screen "Inert Gas Generator Setup" 1280x800, template "Template"
   Circle "Circle_2" at 221,236 size 29x29
      Appearance <- "82_To_HMI_CRNT_MODE_IGG"
   Button "HmiScreenItemData_1" at 1,1 size 150x43; TextOn 'Back'; TextOff 'Main Index'
      on Release: ActivateScreen("02 Main Index", 0)
   Button "HmiScreenItemData_8" at 44,70 size 230x29; TextOn 'Back'; TextOff 'IGGS Mode of Operation'
   Circle "Circle_1" at 221,177 size 29x29
      Appearance <- "82_To_HMI_CRNT_MODE_IGG"
   Button "HmiScreenItemData_4" at 50,167 size 150x51; TextOn 'Back'; TextOff 'Manual'; Authorization "Operate"
      on Press: function_b14e0dd5("80_From_HMI_Request_Manual(1)", 0)
   Circle "Circle_9" at 221,116 size 29x29
      Appearance <- "82_To_HMI_CRNT_MODE_IGG"
   TextField "Text field_1" at 54,547 size 182x20; Text 'Cooling System Overrun'
   TextField "Text field_2" at 54,589 size 192x20; Text 'BWT O2 Content Setpoint'
   TextField "Text field_3" at 54,511 size 89x20; Text 'Description'
   TextField "Text field_5" at 54,670 size 274x20; Text 'IGG Combustion Chamber Post Purge'
   TextField "Text field_6" at 347,511 size 68x20; Text 'Setpoint'
   Button "HmiScreenItemData_6" at 44,467 size 401x29; TextOn 'Back'; TextOff 'IGGS Settings'
   IOField "I/O field_4" at 345,542 size 90x30; Authorization "Commissioning"; FormatPattern 999; Unit  s
      ProcessValue <- "80_From_HMI_Cooling System Overrun"
   IOField "I/O field_5" at 345,583 size 90x30; Authorization "Commissioning"; FormatPattern 99.99; Unit %
      ProcessValue <- "84_Setpoints_E600_BWT_Target"
   IOField "I/O field_6" at 345,664 size 90x30; Authorization "Commissioning"; FormatPattern 999; Unit  s
      ProcessValue <- "80_From_HMI_Post Purge Time"
   TextField "Text field_4" at 54,711 size 294x20; Text 'Air / Inert Gas Pressure (Pre-Ignition)'
   IOField "I/O field_1" at 345,706 size 90x30; Authorization "Commissioning"; FormatPattern 999; Unit  mBar
      ProcessValue <- "84_Setpoints_PIT402_Pilot_Target"
   TextField "Text field_13" at 293,112 size 93x21; Text 'Description'
   IOField "I/O field_13" at 463,150 size 226x30; FormatPattern 9999999999999999999999999999999999999999
      ProcessValue <- "db_time_sync_time_system_READ"
   Button "HmiScreenItemData_26" at 284,70 size 421x29; TextOn 'Back'; TextOff 'Time Setting'
   Button "HmiScreenItemData_24" at 291,192 size 166x30; TextOn 'Back'; TextOff 'Set System Time'; Authorization "Parameter Change"
      on Activate: function_cbf290fd(0, 0)
   Button "HmiScreenItemData_16" at 894,69 size 187x29; TextOn 'Back'; TextOff 'IO'
   Button "HmiScreenItemData_2" at 719,69 size 163x29; TextOn 'Back'; TextOff 'Runtime'
   Button "HmiScreenItemData_10" at 725,107 size 150x51; TextOn 'Back'; TextOff 'Reset AUTO'; Authorization "User administration"
      on Press: function_b14e0dd5("80_From_HMI_RST_AUT_SEQ(1)", 0)
      Appearance <- "80_From_HMI_RST_AUT_SEQ(1)"
   DateTimeField "Date/time field_1" at 463,192 size 226x30; Authorization "Parameter Change"
   TextField "Text field_14" at 314,156 size 142x20; Text 'System Time (UTC)'
   Button "HmiScreenItemData_49" at 44,348 size 401x29; TextOn 'Back'; TextOff 'Inert Gas Transfer Mode'
   Circle "Circle_21" at 400,386 size 26x26
      Appearance <- "80_From_HMI_BWT_BYPASS"
   Button "HmiScreenItemData_50" at 67,384 size 304x33; TextOn 'Back'; TextOff 'Ballast Water Treatment'
      on Press: InvertBit("80_From_HMI_BWT_BYPASS(1)"); ResetBit("80_From_HMI_CRG_BLNK_MODE(1)")
      Appearance <- "80_From_HMI_BWT_BYPASS(1)"
      ObjectEnable <- "100_GCU_AUTO_SEQ_DB_CRNT_STEP"
   Circle "Circle_22" at 400,424 size 26x26
      Appearance <- "80_From_HMI_CRG_BLNK_MODE"
   Button "HmiScreenItemData_51" at 67,422 size 304x33; TextOn 'Back'; TextOff 'Cargo Blanketing'
      on Press: InvertBit("80_From_HMI_CRG_BLNK_MODE(1)"); ResetBit("80_From_HMI_BWT_BYPASS(1)")
      Appearance <- "80_From_HMI_CRG_BLNK_MODE(1)"
      ObjectEnable <- "100_GCU_AUTO_SEQ_DB_CRNT_STEP"
   Button "HmiScreenItemData_23" at 50,106 size 150x51; TextOn 'Back'; TextOff 'Full Automation'; Authorization "Operate"
      on Press: function_b14e0dd5("80_From_HMI_Request_Auto(1)", 0)
   Button "HmiScreenItemData_3" at 1129,1 size 150x43; TextOn 'I&A Compressor Ok'; TextOff 'Back'
      on Release: function_efd93a16()
   IOField "I/O field_2" at 345,747 size 90x30; Authorization "Commissioning"; FormatPattern 999; Unit  mBar
      ProcessValue <- "84_Setpoints_PIT402_Main_Target"
   TextField "Text field_7" at 54,752 size 302x20; Text 'Air / Inert Gas Pressure (Post-Ignition)'
   Button "HmiScreenItemData_7" at 50,228 size 150x51; TextOn 'Back'; TextOff 'FAT Mode'; Authorization "User administration"
      on Press: InvertBit("80_From_HMI_FAT_Mode"); function_b14e0dd5("80_From_HMI_Request_Auto(1)", 0)
   Button "HmiScreenItemData_11" at 725,226 size 150x51; TextOn 'Back'; TextOff 'IGG Standalone'; Authorization "Commissioning"
      on Press: InvertBit("80_From_HMI_IGG_STND_ALN")
      Appearance <- "80_From_HMI_IGG_STND_ALN"
   Button "HmiScreenItemData_12" at 910,107 size 150x35; TextOn 'Back'; TextOff 'P301 Present'; Authorization "Operating Mode"; TextList "P301 Present"
      on Press: InvertBit("80_From_HMI_P301_PRSNT(1)")
      Appearance <- "80_From_HMI_P301_PRSNT(1)"
      ProcessValue <- "80_From_HMI_P301_PRSNT(1)"
   Button "HmiScreenItemData_13" at 910,181 size 150x35; TextOn 'Back'; TextOff 'CV312 Present'; Authorization "User administration"; TextList "CV312 Present"
      on Press: InvertBit("80_From_HMI_CV312_PRSNT")
      Appearance <- "80_From_HMI_CV312_PRSNT"
      ProcessValue <- "80_From_HMI_CV312_PRSNT"
   Button "HmiScreenItemData_14" at 910,218 size 150x35; TextOn 'Back'; TextOff 'CV431 Present'; Authorization "Operating Mode"; TextList "CV431 Present"
      on Press: InvertBit("80_From_HMI_CV431_PRSNT")
      Appearance <- "80_From_HMI_CV431_PRSNT"
      ProcessValue <- "80_From_HMI_CV431_PRSNT"
   Button "HmiScreenItemData_15" at 910,255 size 150x35; TextOn 'Back'; TextOff 'CV432 Present'; Authorization "Operating Mode"; TextList "CV432 Present"
      on Press: InvertBit("80_From_HMI_CV432_PRSNT")
      Appearance <- "80_From_HMI_CV432_PRSNT"
      ProcessValue <- "80_From_HMI_CV432_PRSNT"
   Button "HmiScreenItemData_18" at 725,166 size 150x51; TextOn 'Back'; TextOff 'Silence Buzzer'; Authorization "Operate"
      on Press: function_b14e0dd5("80_From_HMI_SLNCE_BZR", 0)
      Appearance <- "80_From_HMI_SLNCE_BZR"
   IOField "I/O field_7" at 596,369 size 93x43; Authorization "Commissioning"; FormatPattern 999; Unit  step
      ProcessValue <- "100_IGG_AUTO_SEQ_DB_CRNT_STEP"
   IOField "I/O field_8" at 598,426 size 93x43; Authorization "Commissioning"; FormatPattern 999; Unit  step
      ProcessValue <- "100_BC_AUTO_SEQ_DB_CRNT_STEP"
   Button "HmiScreenItemData_9" at 485,376 size 102x29; TextOn 'Back'; TextOff 'IGG PLC'
   Button "HmiScreenItemData_17" at 485,433 size 102x29; TextOn 'Back'; TextOff 'BC PLC'
   Button "HmiScreenItemData_19" at 700,376 size 563x29; TextOn 'Back'; TextOff 'IGG STEP'; TextList "STEP LIST IGG"
      ProcessValue <- "100_IGG_AUTO_SEQ_DB_CRNT_STEP"
   Button "HmiScreenItemData_20" at 700,433 size 563x29; TextOn 'Back'; TextOff 'IGG STEP'; TextList "STEP LIST BC"
      ProcessValue <- "100_BC_AUTO_SEQ_DB_CRNT_STEP"
   AlarmView "Alarm view_1" at 0,777 size 1280x23
   IOField "I/O field_9" at 618,295 size 60x30; Authorization "Operate"; FormatPattern 99; Unit  s
      ProcessValue <- "80_From_HMI_Beacon frequency"
   IOField "I/O field_10" at 619,332 size 60x30; Authorization "Operate"; FormatPattern 99; Unit  min
      ProcessValue <- "80_From_HMI_Buzzer reset time"
   TextField "Text field_9" at 489,301 size 138x20; Text 'Beacon frequency'
   TextField "Text field_10" at 489,337 size 100x20; Text 'Buzzer reset'
   TextField "Text field_11" at 974,670 size 257x27; Text 'Proportionate Component PID'
   TextField "Text field_15" at 974,704 size 257x27; Text 'Integrative Component PID'
   TextField "Text field_16" at 974,737 size 257x27; Text 'Derivative Component PID'
   TextField "Text field_17" at 976,486 size 153x27; Text 'GAIN'
   TextField "Text field_18" at 974,515 size 153x27; Text 'Integration Time'
   TextField "Text field_19" at 974,549 size 153x27; Text 'Derivation Time'
   TextField "Text field_20" at 976,584 size 153x27; Text 'Maximum opening'
   Group "Group_15" at 1129,515 size 112x34; Authorization "User administration"; Picture "Graphic_284"; FormatPattern 99
   Group "Group_16" at 1129,550 size 112x34; Authorization "User administration"; Picture "Graphic_284"; FormatPattern 99
   Group "Group_3" at 1129,480 size 112x34; Authorization "User administration"; Picture "Graphic_284"; FormatPattern 99
   Switch "Switch_8" at 1222,670 size 32x29; CaptionText 'Switch'; TextOn 'ON'; TextOff 'OFF'; Authorization "User administration"; PictureOff "Design_5_PilotLight_Green_Off"; PictureOn "Design_5_PilotLight_Green_On"
      on Change: InvertBit("84_Setpoints_P_ON")
      ProcessValue <- "84_Setpoints_P_ON"
   Switch "Switch_9" at 1222,704 size 32x29; CaptionText 'Switch'; TextOn 'ON'; TextOff 'OFF'; Authorization "User administration"; PictureOff "Design_5_PilotLight_Green_Off"; PictureOn "Design_5_PilotLight_Green_On"
      on Change: InvertBit("84_Setpoints_I_ON")
      ProcessValue <- "84_Setpoints_I_ON"
   Switch "Switch_10" at 1222,735 size 32x29; CaptionText 'Switch'; TextOn 'ON'; TextOff 'OFF'; Authorization "User administration"; PictureOff "Design_5_PilotLight_Green_Off"; PictureOn "Design_5_PilotLight_Green_On"
      on Change: InvertBit("84_Setpoints_D_ON")
      ProcessValue <- "84_Setpoints_D_ON"
   Group "Group_1" at 1129,618 size 112x34; Picture "Graphic_284"; Authorization "Commissioning"; FormatPattern 99
   TextField "Text field_21" at 976,618 size 153x27; Text 'Minimum opening'
   Gauge "Gauge_1" at 699,468 size 239x239; UnitText '%'; CaptionText 'CV 203'
      ProcessValue <- "16_AQ_Data_CV203_CNTRL"
   Circle "Circle_29" at 707,748 size 20x20
      Appearance <- "Evolving Setpoint_DB_LevelBetter"
   TextField "Text field_22" at 736,744 size 199x27; Text 'O2 content geting Better'
   Gauge "Gauge_2" at 456,468 size 239x239; UnitText '%'; CaptionText 'O2 Content'
      Visibility <- "80_From_HMI_CRG_BLNK_MODE"
      ProcessValue <- "12_AI_Data_E600O2ContentIn"
      MaximumValue <- "84_Setpoints_E600_CB_HighHigh"
   Button "Button_25" at 582,743 size 95x31; TextOn 'grafic'; TextOff 'GRAFIC'; PictureOff "imageedit_175_8204096749"
      on Click: function_efd93a16("CV 203 Grafics", 200, 100, -1, -1, 1)
   Gauge "Gauge_3" at 456,468 size 239x239; UnitText '%'; CaptionText 'O2 Content'
      Visibility <- "80_From_HMI_BWT_BYPASS"
      ProcessValue <- "12_AI_Data_E600O2ContentIn"
      MaximumValue <- "84_Setpoints_E600_BWT_HighHigh"
   Group "Group_2" at 1129,584 size 112x34; Picture "Graphic_284"; Authorization "Commissioning"; FormatPattern 99
   Button "HmiScreenItemData_21" at 910,144 size 150x35; TextOn 'Back'; TextOff 'P305 Present'; Authorization "Operating Mode"; TextList "P305 Present"
      on Press: InvertBit("80_From_HMI_P305_PRSNT")
      Appearance <- "80_From_HMI_P305_PRSNT"
      ProcessValue <- "80_From_HMI_P305_PRSNT"
   TextField "Text field_8" at 54,630 size 154x20; Text 'Cargo Blanketing O2'
   IOField "I/O field_3" at 345,624 size 90x30; Authorization "Commissioning"; FormatPattern 99.99; Unit %
      ProcessValue <- "84_Setpoints_E600_CB_Target"
   GraphicView "Graphic view_22" at 1129,515 size 112x34; Picture "Graphic_284"
   IOField "D5_I/O field_2" at 1144,523 size 62x18; Authorization "User administration"; FormatPattern 99999
      ProcessValue <- "84_Setpoints_Integration Time"
   TextField "D5_Text field_2" at 1204,523 size 23x18; Text 'ms / km/h'
   GraphicView "Graphic view_23" at 1129,550 size 112x34; Picture "Graphic_284"
   IOField "D5_I/O field_3" at 1144,558 size 62x18; FormatPattern 99999
      ProcessValue <- "84_Setpoints_Derive Time"
   TextField "D5_Text field_3" at 1204,558 size 23x18; Text 'ms / km/h'
   GraphicView "Graphic view_25" at 1129,480 size 112x34; Picture "Graphic_284"
   IOField "D5_I/O field_10" at 1144,488 size 62x18; Authorization "User administration"; FormatPattern 99.9999
      ProcessValue <- "84_Setpoints_Gain"
   TextField "D5_Text field_10" at 1204,488 size 23x18; Text 'km/h'
   GraphicView "Graphic view_1" at 1129,618 size 112x34; Picture "Graphic_284"
   IOField "D5_I/O field_1" at 1144,626 size 62x18; Authorization "Commissioning"; FormatPattern 999
      ProcessValue <- "84_Setpoints_Min Opening"
   TextField "D5_Text field_1" at 1204,626 size 23x18; Text '% / km/h'
   GraphicView "Graphic view_2" at 1129,584 size 112x34; Picture "Graphic_284"
   IOField "D5_I/O field_5" at 1144,592 size 62x18; Authorization "Commissioning"; FormatPattern 999
      ProcessValue <- "84_Setpoints_Max Opening"
   TextField "D5_Text field_5" at 1204,592 size 23x18; Text '% / km/h'

screen "Reports" 1280x800, template "Template"
   RecipeView "Recipe view_1" at 854,43 size 400x365; Tag4DataRecord "Record Data Tag"; Tag4RecipeNumber "Recipe Tag"
   Button "HmiScreenItemData_1" at 2,2 size 159x51; TextOn 'Back'; TextOff 'Home'
      on Release: ActivateScreen("01 Home", 0)

PopupScreen "BWT Mode Warning" 665x250
   Button "Button_1" at 0,0 size 665x250; TextOff 'BWT Mode Not Selected. Select BWT Mode for Tank Treatment. For Cargo Blanketing use IGG Controls.'
      on Release: ActivateScreen("Balast Water Treatment Setup", 0)
   Button "Button_2" at 208,187 size 250x35; TextOff 'OK, Select Treatment Mode'
      on Release: ActivateScreen("Balast Water Treatment Setup", 0); function_efd93a16("BWT Mode Warning", 0, 0, -1, -1, 1)

PopupScreen "CV 203 Grafics" 810x675
   Button "Button_1" at 753,0 size 56x38; TextOff 'Text'; PictureOff "Graphic_286"
      on Click: function_efd93a16("CV 203 Grafics", 0, 0, -1, -1, 1)
   GraphicView "Graphic view_2" at 2,2 size 751x35; Picture "Graphic_287"
   TextField "Text field_1" at 285,7 size 229x26; Text 'O2 FUEL MODULATION'
   TrendView "Trend view_2" at 1,38 size 808x636
      Visibility <- "80_From_HMI_CRG_BLNK_MODE"
      ValueAxis2End <- "84_Setpoints_Max Opening"
      ValueAxis2Begin <- "84_Setpoints_Min Opening"
      ValueAxis1End <- "84_Setpoints_E600_CB_HighHigh"
   TrendView "Trend view_1" at 2,40 size 804x635
      Visibility <- "80_From_HMI_BWT_BYPASS"
      ValueAxis2End <- "84_Setpoints_Max Opening"
      ValueAxis2Begin <- "84_Setpoints_Min Opening"
      ValueAxis1End <- "84_Setpoints_E600_BWT_HighHigh"

PopupScreen "CV 403 Grafics" 810x675
   Button "Button_1" at 753,0 size 56x40; TextOff 'Text'; PictureOff "Graphic_286"
      on Click: function_efd93a16("CV 403 Grafics", 0, 0, -1, -1, 1)
   GraphicView "Graphic view_2" at 2,2 size 751x35; Picture "Graphic_287"
   TextField "Text field_1" at 285,9 size 281x26; Text 'IG PRESSURE MODULATION'
   TrendView "Trend view_2" at 1,39 size 809x635

PopupScreen "Double Block & Bleed Valve Monitoring" 497x370
   Button "Button_1" at 3,1 size 490x365; TextOff 'Text'
      on Release: function_efd93a16("Double Block & Bleed Valve Monitoring", 250, 250, -1, -1, 1)
   GraphicView "Graphic view_59" at 119,276 size 259x20; Picture "Graphic_151"
   Group "Group_2" at 159,200 size 58x100; Picture "Graphic_72"
   TextField "Text field_45" at 159,219 size 54x20; Text 'Closed'
      Visibility <- "10_DI_DATA_CV407_CLSD"
   GraphicView "Graphic view_58" at 237,172 size 19x110; Picture "Graphic_147"
   GraphicView "Graphic view_60" at 233,145 size 58x58; Picture "Graphic_162"
   TextField "Text field_6" at 148,304 size 80x22; Text 'CV407'
   TextField "Text field_8" at 269,304 size 79x22; Text 'CV411'
   Group "Group_3" at 279,200 size 58x100; Picture "Graphic_72"
   GraphicView "Graphic view_65" at 237,138 size 19x21; Picture "Graphic_147"
   TextField "Text field_9" at 281,219 size 54x20; Text 'Closed'
      Visibility <- "10_DI_DATA_CV411_CLSD"
   TextField "Text field_10" at 281,219 size 54x20; Text 'Opened'
      Visibility <- "10_DI_DATA_CV411_OPN"
   TextField "Text field_12" at 290,165 size 54x20; Text 'Closed'
      Visibility <- "10_DI_DATA_CV409_CLSD"
   TextField "Text field_13" at 290,165 size 54x20; Text 'Opened'
      Visibility <- "10_DI_DATA_CV409_OPN"
   TextField "Text field_5" at 244,117 size 75x22; Text 'CV409'
   Circle "Circle_28" at 266,282 size 10x10
      Visibility <- "10_DI_DATA_CV407_OPN"
   Circle "Circle_29" at 215,282 size 10x10
      Visibility <- "10_DI_DATA_CV407_OPN"
   Circle "Circle_30" at 337,282 size 10x10
      Visibility <- "10_DI_DATA_CV411_OPN"
   TextField "Text field_11" at 159,219 size 54x20; Text 'Opened'
      Visibility <- "10_DI_DATA_CV407_OPN"
   Circle "Circle_42" at 244,280 size 10x10
      Visibility <- "10_DI_DATA_CV407_OPN"
   Circle "Circle_43" at 359,278 size 10x10
      Visibility <- "10_DI_DATA_CV411_OPN"
   Circle "Circle_44" at 242,204 size 10x10
      Visibility <- "10_DI_DATA_CV409_OPN"
   TextField "Text field_1" at 85,79 size 327x30; Text 'Double Block & Bleed Valves'
   Button "Button_2" at 10,10 size 109x40; TextOff 'DB&B'
      on Release: function_efd93a16("Double Block & Bleed Valve Monitoring", 250, 250, -1, -1, 1)
   Circle "Circle_1" at 242,234 size 10x10
      Visibility <- "10_DI_DATA_CV409_OPN"
   Circle "Circle_2" at 149,281 size 10x10
      Visibility <- "10_DI_DATA_CV407_OPN"
   GraphicView "Graphic view_63" at 159,200 size 58x100; Picture "Graphic_72"
   GraphicView "Graphic view_64" at 279,200 size 58x100; Picture "Graphic_72"

PopupScreen "IGG Temperature Trends" 810x675
   on GenerateScreen: "TitleUpdater"()
   Button "Button_1" at 753,0 size 56x38; TextOff 'Text'; PictureOff "Graphic_286"
      on Click: function_efd93a16("IGG Temperature Trends", 0, 0, -1, -1, 1)
   GraphicView "Graphic view_2" at 2,2 size 751x35; Picture "Graphic_287"
   TrendView "Trend view_1" at 1,40 size 805x635
      Visibility <- "80_From_HMI_BWT_BYPASS"
      ValueAxis2End <- "84_Setpoints_PIT359_HighHigh"
      ValueAxis2Begin <- "84_Setpoints_PIT359_LowLow"
   TextField "Text field_1" at 282,7 size 252x26; Text 'IGG Temperature Trends'

PopupScreen "PGC Commissioning" 1280x800
   Button "Button_1" at 308,285 size 665x230; TextOff 'Text'
      on Release: ActivateScreen("Inert Gas Generator Plant", 0)
   Button "Button_2" at 540,431 size 200x55; TextOff 'OK'
      on Release: ResetBit("PGC_COMMISSION_MODE_DB_Active")
   TextField "Text field_1" at 303,313 size 674x100; Text 'Tanks can now be changed over, press OK when completed'

PopupScreen "Salinity - Acceptance" 1050x350
   Button "Button_2" at 556,290 size 105x50; TextOff 'NO'
      on Release: ActivateScreen("Balast Water Treatment Setup", 0)
   Button "Button_3" at 390,290 size 105x50; TextOff 'YES'
      on Press: function_b14e0dd5("80_From_HMI_SAL_CNFRM", 0)
      on Release: function_efd93a16("Salinity - Acceptance", 168, 315, -1, -1, 1)
   TextField "Text field_1" at 223,102 size 604x82; Text 'Please confirm that the entered salinity value of is correct'
   IOField "I/O field_1" at 510,138 size 139x50; FormatPattern 99.9; Unit  psu
      ProcessValue <- "80_From_HMI_SAL_VALUE"

PopupScreen "Salinity - Fresh Water Alert" 1280x800
   Button "Button_1" at 115,225 size 1050x284; TextOff 'NOTE: BALLAST WATER SALINITY IS FRESH WATER LEVEL This System Is Not Certified For FRESH WATER Treatment. Do Wish To Continue Ballast Water Treatment?'
   Button "Button_2" at 666,514 size 105x50; TextOff 'NO'
      on Release: ActivateScreen("Balast Water Treatment Setup", 0)
      on Press: function_b14e0dd5("80_From_HMI_LOW_SAL_RJCT", 0)
   Button "Button_3" at 500,514 size 105x50; TextOff 'YES'
      on Release: ActivateScreen("Balast Water Treatment Setup", 0)
      on Press: function_b14e0dd5("80_From_HMI_LOW_SAL_ACPT", 0)

PopupScreen "SD Card overflow" 665x230
   Button "Button_1" at 0,0 size 665x230; TextOff 'Data Logging SD Card Memory Full'
      on Click: function_efd93a16("SD Card overflow", 0, 0, -1, -1, 1)
      on Press: ResetBit("Logging SD Card Overflow")

PopupScreen "Start Treatment" 665x230
   Button "Button_1" at 0,0 size 665x230; TextOff 'Text'
   Button "Button_2" at 232,146 size 200x55; TextOff 'OK'; Authorization "Operate"
      on Release: function_efd93a16("Start Treatment", 0, 0, -1, -1, 1); ActivateScreen("Inert Gas Generator Plant", 0)
   TextField "Text field_1" at 72,25 size 520x52; Text 'Treatment now required'
   TextField "Text field_2" at 16,75 size 644x64; Text 'Please Make Sure the Energy and Water Supply are Present and Sufficient'

PopupScreen "Time Until Treatment Required" 750x270
   Button "Button_1" at 0,0 size 750x270; TextOff 'Text'
   Button "Button_2" at 268,157 size 200x55; TextOff 'OK'; Authorization "Operate"
      on Click: function_efd93a16("Time Until Treatment Required", 0, 0, -1, -1, 1); ActivateScreen("Inert Gas Generator Plant", 0)
   TextField "Text field_1" at 6,24 size 728x100; Text 'Treatment required to start in hours and minutes'
   IOField "I/O field_1" at 207,72 size 104x52; FormatPattern 99
      ProcessValue <- "Sequence Times_DB_Pre-Dwell Timer_Hours Left"
   IOField "I/O field_2" at 470,72 size 104x52; FormatPattern 99
      ProcessValue <- "Sequence Times_DB_Pre-Dwell Timer_Minutes Left"

PopupScreen "Treatment check / Daily Checks Completed" 1050x350
   Button "Button_3" at 411,283 size 229x50; TextOff 'CONFIRM'
      on Release: function_efd93a16("Treatment check / Daily Checks Completed", 0, 0, 0, -1, 1)
      on Press: function_b14e0dd5("88_treatment_POP_UP_CNFRM", 0)
   TextField "Text field_1" at 3,36 size 1044x240; Text 'Please confirm pre treatment check and daily checks are completed.'

PopupScreen "Treatment Cycle Completed" 665x230
   Button "Button_1" at 0,0 size 665x230; TextOff 'TREATMENT CYCLE COMPLETED'
      on Click: function_efd93a16("Treatment Cycle Completed", 0, 0, -1, -1, 1)

PopupScreen "Treatment Status" 300x280
   Button "HmiScreenItemData_40" at 0,0 size 300x29; TextOn 'Back'; TextOff 'Treatment Status'
      on Release: function_efd93a16("Treatment Status", 0, 0, -1, -1, 1)
   Button "HmiScreenItemData_9" at 17,34 size 220x30; TextOn 'Back'; TextOff 'Pre Dwell Time Completed'
      on Release: function_efd93a16("Treatment Status", 0, 0, -1, -1, 1)
   Button "HmiScreenItemData_17" at 17,94 size 220x30; TextOn 'Back'; TextOff 'De-Oxygenation Completed'
      on Release: function_efd93a16("Treatment Status", 0, 0, -1, -1, 1)
   Button "HmiScreenItemData_38" at 17,124 size 220x30; TextOn 'Back'; TextOff 'Dwell Time Completed'
      on Release: function_efd93a16("Treatment Status", 0, 0, -1, -1, 1)
   Button "HmiScreenItemData_39" at 17,184 size 220x30; TextOn 'Back'; TextOff 'Re-Oxygenation Completed'
      on Release: function_efd93a16("Treatment Status", 0, 0, -1, -1, 1)
   Button "HmiScreenItemData_41" at 18,215 size 220x30; TextOn 'Back'; TextOff 'Post Dwell Time Completed'
      on Release: function_efd93a16("Treatment Status", 0, 0, -1, -1, 1)
   Button "HmiScreenItemData_46" at 17,64 size 220x30; TextOn 'Back'; TextOff 'Inert Gas Transfer Active'
   Button "HmiScreenItemData_48" at 17,154 size 220x30; TextOn 'Back'; TextOff 'Ambient Air Transfer Active'
   Button "HmiScreenItemData_52" at 17,64 size 220x30; TextOn 'Back'; TextOff 'IG Transfer Completed'
      on Release: function_efd93a16("Treatment Status", 0, 0, -1, -1, 1)
   Button "HmiScreenItemData_53" at 17,154 size 220x30; TextOn 'Back'; TextOff 'Ambient Air Transfer Completed'
      on Release: function_efd93a16("Treatment Status", 0, 0, -1, -1, 1)
   Button "Button_2" at 0,0 size 34x29; TextOff 'Text'; PictureOff "Graphic_286"
      on Click: function_efd93a16("Treatment Status", 0, 0, -1, -1, 1)
   Circle "Circle_23" at 254,38 size 24x24
      Appearance <- "2110_BTCS_CNTRL_DB_BTCS_STEP"
   Circle "Circle_24" at 254,67 size 24x24
      Appearance <- "100_GCU_AUTO_SEQ_DB_CRNT_STEP"
   Circle "Circle_25" at 254,97 size 24x24
      Appearance <- "2110_BTCS_CNTRL_DB_BTCS_STEP"
   Circle "Circle_26" at 254,127 size 24x24
      Appearance <- "2110_BTCS_CNTRL_DB_BTCS_STEP"
   Circle "Circle_27" at 254,157 size 24x24
      Appearance <- "100_GCU_AUTO_SEQ_DB_CRNT_STEP"
   Circle "Circle_28" at 254,187 size 24x24
      Appearance <- "2110_BTCS_CNTRL_DB_BTCS_STEP"
   Circle "Circle_29" at 254,217 size 24x24
      Appearance <- "2110_BTCS_CNTRL_DB_BTCS_STEP"

PopupScreen "Voyage Time Warning" 665x250
   Button "Button_1" at 0,0 size 665x250; TextOff 'Voyage Time Insufficient, Minimum Voyage Time For Treatment Is Days.'
      on Release: ActivateScreen("Balast Water Treatment Setup", 0)
   IOField "I/O field_1" at 359,124 size 82x50; FormatPattern 999
      ProcessValue <- "2102_TIME_CALCS_DB_TOT_SEQ_DAYS"
   Button "Button_2" at 208,187 size 250x35; TextOff 'OK, Adjust Voyage Time'
      on Release: ActivateScreen("Balast Water Treatment Setup", 0); function_efd93a16("Voyage Time Warning", 0, 0, -1, -1, 1)

screen "02 Main Index" 1280x800, template "Template"
   on GenerateScreen: "User_Change"()
   GraphicView "Graphic view_1" at 314,58 size 650x705; Picture "Graphic_115"
   TextField "HmiScreenItemData_16" at 80,95 size 880x30; Text 'BALLAST WATER MANAGEMENT SYSTEM'
   Button "HmiScreenItemData_17" at 320,150 size 160x60; TextOn 'IGG Plant'; TextOff 'IGG Plant'; Authorization "Operate"
      on Release: ActivateScreen("Inert Gas Generator Plant", 0)
   Button "HmiScreenItemData_20" at 800,250 size 160x60; TextOn 'IGG Plant'; TextOff 'Commissioning'; Authorization "Commissioning"
      on Release: ActivateScreen("Commissioning Main Page", 0)
   Button "HmiScreenItemData_1" at 2,2 size 159x51; TextOn 'Back'; TextOff 'Home'
      on Release: ActivateScreen("01 Home", 0)
   Button "HmiScreenItemData_4" at 560,250 size 160x60; TextOn 'IGG Plant'; TextOff 'Air System'; Authorization "Operate"
      on Release: ActivateScreen("Air System", 0)
   Button "HmiScreenItemData_7" at 560,150 size 160x60; TextOn 'IGG Plant'; TextOff 'Fuel System'; Authorization "Operate"
      on Release: ActivateScreen("Fuel System", 0)
   Button "HmiScreenItemData_5" at 80,150 size 160x60; TextOn 'IGG Plant'; TextOff 'IGG Setup'; Authorization "Commissioning"
      on Release: ActivateScreen("Inert Gas Generator Setup", 0)
   Button "Button_1" at 800,650 size 160x60; TextOn 'User Account'; TextOff 'User Administration'; Authorization "User administration"
      on Release: ActivateScreen("03 User Admin", 0)
   Button "HmiScreenItemData_9" at 1147,54 size 125x51; TextOn 'IGG Plant'; TextOff 'Login'
      on Click: function_a2a04561()
      on Release: ActivateScreen("Commissioning Main Page", 0)
   Button "HmiScreenItemData_12" at 1147,2 size 125x51; TextOn 'IGG Plant'; TextOff 'Logout'
      on Release: function_f23ef4c9()
   IOField "I/O field_1" at 991,137 size 266x35; FormatPattern ???????????????????????
      ProcessValue <- "Current User"
   Button "HmiScreenItemData_13" at 560,450 size 160x60; TextOn 'IGG Plant'; TextOff 'Fresh Water System'; Authorization "Operate"
      on Release: ActivateScreen("Fresh Water System", 0)
   Button "HmiScreenItemData_2" at 560,350 size 160x60; TextOn 'IGG Plant'; TextOff 'Cooling System'; Authorization "Operate"
      on Release: ActivateScreen("Cooling System", 0)
   Button "Button_2" at 800,150 size 160x60; TextOn 'User Account'; TextOff 'Alarm Log'; Authorization "Operate"
      on Release: ActivateScreen("04 Alarm Log", 0)
   Button "HmiScreenItemData_6" at 320,250 size 160x60; TextOn 'IGG Plant'; TextOff 'GCU Plant'; Authorization "Operate"
      on Release: ActivateScreen("Inert Gas Conditioning Plant", 0)
   Button "HmiScreenItemData_8" at 80,250 size 160x60; TextOn 'IGG Plant'; TextOff 'GCU Setup'; Authorization "Commissioning"
      on Release: ActivateScreen("Inert Gas Conditioning Setup", 0)
   Button "HmiScreenItemData_10" at 320,350 size 160x60; TextOn 'IGG Plant'; TextOff 'BWT Plant'; Authorization "Operate"
      on Release: ActivateScreen("Balast Water Treatment Plant", 0)
   Button "HmiScreenItemData_11" at 91,575 size 160x60; TextOn 'IGG Plant'; TextOff 'BWT Setup'; Authorization "Operate"
      on Release: ActivateScreen("42 BWT Setup", 0)
      Visibility <- "AlwaysTRUE"
   Button "Button_3" at 560,550 size 160x60; TextOn 'User Account'; TextOff 'IG Transfer Mode'; Authorization "Operate"
      on Release: ActivateScreen("IG Transfer Mode", 0)
   Button "Button_4" at 91,455 size 160x60; TextOn 'User Account'; TextOff 'BTCS Setup & Launch'; Authorization "User administration"
      on Release: ActivateScreen("08 BTCS MAIN", 0)
      Visibility <- "AlwaysTRUE"
   Button "Button_5" at 800,350 size 160x60; TextOn 'User Account'; TextOff 'System Configuration'; Authorization "Commissioning"
      on Release: ActivateScreen("09 Sys Config", 0)
   Button "Button_6" at 80,650 size 400x60; TextOn 'User Account'; TextOff 'BWTS (Balast Water Treatment System) Setup & Launch'; Authorization "User administration"
      on Release: ActivateScreen("07 BWTS MAIN", 0)
      Visibility <- "AlwaysTRUE"
   Button "Button_7" at 560,650 size 160x60; TextOn 'User Account'; TextOff 'PGC System'; Authorization "Operate"
      on Release: ActivateScreen("PGC System", 0)
   Button "Button_8" at 60,411 size 200x29; TextOn 'User Account'; TextOff 'Tank Control System'; Authorization "User administration"
   Button "Button_9" at 80,350 size 160x60; TextOn 'User Account'; TextOff 'BTCS Setup & Launch'; Authorization "Operate"
      on Release: ActivateScreen("Balast Water Treatment Setup", 0)
   Button "Button_10" at 800,450 size 160x60; TextOn 'User Account'; TextOff 'Report Test'; Authorization "User administration"
      on Release: ActivateScreen("Reports", 0)
      Visibility <- "user_group"

screen "Balast Water Treatment Plant Tank Levels" 1280x800, template "Template"
   on GenerateScreen: "User_Change"(); "TitleUpdater"()
   Button "HmiScreenItemData_1" at 1,1 size 150x40; TextOn 'Back'; TextOff 'Main Index'
      on Release: ActivateScreen("02 Main Index", 0)
   TextField "Text field_63" at 383,107 size 72x30; Text 'Pre Dwell Time'
   Circle "Circle_29" at 1047,85 size 20x20
      Appearance <- "2102_TIME_CALCS_DB_POST_DWELL_TMR_DN"
   Button "HmiScreenItemData_9" at 10,60 size 158x27; TextOn 'Back'; TextOff 'BWTS Control'
   Button "HmiScreenItemData_4" at 14,150 size 75x47; TextOn 'Back'; TextOff 'Stop'; Authorization "Operate"
      ObjectEnable <- "82_To_HMI_CRNT_MODE_GCU"
      on Release: function_efd93a16("BWTS Stop Confirm", 400, 200, -1, -1, 1)
   Circle "Circle_20" at 137,105 size 29x29
      Appearance <- "82_To_HMI_IGG RUN Indication"
   Button "HmiScreenItemData_3" at 14,93 size 75x47; TextOn 'Back'; TextOff 'Start'; Authorization "Operate"
      on Release: function_efd93a16("BWTS Start Confirm", 400, 200, -1, -1, 1)
      ObjectEnable <- "82_To_HMI_CRNT_MODE_GCU"
   Button "HmiScreenItemData_2" at 1129,1 size 150x40; TextOn 'Back'; TextOff 'BWTS Setup'
      on Release: ActivateScreen("Balast Water Treatment Setup", 0)
   TextField "Text field_1" at 290,107 size 68x30; Text 'Tank Selected'
   TextField "Text field_2" at 841,107 size 61x30; Text 'BWTS Started'
   TextField "Text field_3" at 568,107 size 62x30; Text 'IGGS Started'
   TextField "Text field_4" at 659,107 size 60x30; Text 'GCU Started'
   TextField "Text field_5" at 748,107 size 61x30; Text 'PGC Started'
   TextField "Text field_6" at 908,107 size 102x30; Text 'Gas Transfer Started'
   Circle "Circle_10" at 956,89 size 14x14
      Appearance <- "2110_BTCS_CNTRL_DB_BTCS_STEP"
   TextField "Text field_7" at 995,107 size 125x30; Text 'Treatment Cycle Completed'
   TextField "Text field_23" at 261,291 size 34x14; Text 'MBG'
   GraphicView "Graphic view_17" at 575,446 size 532x12; Picture "Graphic_151"
   Button "Button_13" at 252,437 size 37x30; TextOff 'DB&B'
   TextField "Text field_58" at 188,226 size 50x40; Text 'Safe Area'
   Button "Button_20" at 724,152 size 115x34; TextOff 'Re-Oxygenation'
      Appearance <- "2110_BTCS_CNTRL_DB_BTCS_STEP"
   Button "Button_21" at 845,152 size 93x34; TextOff 'Post Dwell'
      Appearance <- "2110_BTCS_CNTRL_DB_BTCS_STATE"
   Circle "Circle_1" at 137,105 size 29x29
      Appearance <- "2110_BTCS_CNTRL_DB_BTCS_STATE"
   Circle "Circle_8" at 775,89 size 14x14
      Appearance <- "2110_BTCS_CNTRL_DB_BTCS_STEP"
   Circle "Circle_9" at 685,89 size 14x14
      Appearance <- "100_GCU_AUTO_SEQ_DB_CRNT_STEP"
   Circle "Circle_11" at 595,89 size 14x14
      Appearance <- "51_SLAVE_STATUS_RUNNING"
   Circle "Circle_12" at 866,89 size 14x14
      Appearance <- "2110_BTCS_CNTRL_DB_BTCS_STEP"
   Circle "Circle_13" at 324,89 size 14x14
      Appearance <- "HMI Indication Logic_DB_Tank Selected"
   Circle "Circle_14" at 414,89 size 14x14
      Appearance <- "2102_TIME_CALCS_DB_PRE_DWELL_TMR_DN"
   Button "Button_3" at 626,152 size 93x34; TextOff 'Dwell'
      Appearance <- "2110_BTCS_CNTRL_DB_BTCS_STATE"
   Button "Button_5" at 944,152 size 93x34; TextOff 'Complete'
      Appearance <- "HMI Indication Logic_DB_Sequence Finished"
   TextField "Text field_61" at 202,107 size 71x30; Text 'FA Mode Selected'
   Circle "Circle_2" at 230,89 size 14x14
      Appearance <- "HMI Indication Logic_DB_FA Mode Selected"
   TextField "Text field_60" at 190,519 size 46x25; Text 'GCU'
   GraphicIOField "Graphic I/O field_4" at 187,543 size 53x55; PictureList "GCU"
      ProcessValue <- "100_GCU_AUTO_SEQ_DB_RNG"
   TextField "Text field_74" at 186,279 size 54x25; Text 'IGGS'
   GraphicIOField "Graphic I/O field_1" at 185,303 size 57x53; PictureList "IGGS"
      ProcessValue <- "14_DQ_Data_24PF1"
   TextField "Text field_62" at 183,359 size 60x20; Text 'Disabled'
   TextField "Text field_77" at 183,359 size 60x20; Text 'Enabled'
      Visibility <- "51_SLAVE_STATUS_RUNNING"
   Button "Button_8" at 178,280 size 70x105; TextOff 'Text'
      on Release: ActivateScreen("Inert Gas Generator Plant", 0)
   TextField "Text field_70" at 183,599 size 60x20; Text 'Disabled'
   TextField "Text field_71" at 183,599 size 60x20; Text 'Enabled'
      Visibility <- "100_GCU_AUTO_SEQ_DB_RNG"
   Button "Button_4" at 178,521 size 70x105; TextOff 'Text'
      on Release: ActivateScreen("Inert Gas Conditioning Plant", 0)
   GraphicIOField "Graphic I/O field_2" at 770,45 size 250x30; PictureList "Process time Banner"
      ProcessValue <- "2110_BTCS_CNTRL_DB_BTCS_STATE"
      Visibility <- "2110_BTCS_CNTRL_DB_BTCS_STATE"
   Button "Button_14" at 303,152 size 93x34; TextOff 'Unselected'
      Visibility <- "HMI Indication Logic_DB_Tank Selected"
      Appearance <- "HMI Indication Logic_DB_Tank Selected"
   Button "Button_15" at 404,152 size 93x34; TextOff 'Selected'
      Appearance <- "HMI Indication Logic_DB_Tank Selected"
   Button "Button_16" at 506,152 size 115x34; TextOff 'De-Oxygenation'
      Appearance <- "2110_BTCS_CNTRL_DB_BTCS_STEP"
   TextField "Text field_92" at 304,351 size 76x15; Text 'FIT-418-6P'
   TextField "Text field_98" at 304,308 size 76x15; Text 'FIT-420-6P'
   Button "HmiScreenItemData_19" at 1185,676 size 72x27; TextOn 'Back'; TextOff 'Status'
      on Press: function_efd93a16("Treatment Status", 100, 471, -1, 3, 1)
   Group "Group_5" at 664,46 size 45x27; FormatPattern 999
   Group "Group_6" at 298,44 size 241x30
   Circle "Circle_26" at 504,89 size 14x14
      Appearance <- "2102_TIME_CALCS_DB_Time_To_Treatment"
   TextField "Text field_134" at 470,107 size 75x30; Text 'Wait for IGGS Start'
   GraphicView "Graphic view_4" at 357,210 size 25x62; Picture "Graphic_183"
   GraphicView "Graphic view_5" at 265,210 size 25x62; Picture "Graphic_183"
   IOField "I/O field_31" at 1053,45 size 225x30; FormatPattern ???????????????
      ProcessValue <- "Current User"
   Button "HmiScreenItemData_8" at 772,732 size 503x40; TextOn 'Back'; TextOff 'Text'
   TextField "Screen title" at 783,728 size 496x50; Text 'Screen title'
   Bar "Bar_1" at 262,206 size 122x241; MinimumValue 0; MaximumValue 100
      ProcessValue <- "20_TANKS_IP_DATA_RIO_06_FIRST_TANK_BWT_LEVEL"
   Button "Button_48" at 273,396 size 100x25; TextOff 'DISABLED'
      on Release: function_efd93a16("Tank 6P Status", 168, 315, -1, 2, 1)
      Visibility <- "504_Tank Grouping_DB2020_GROUP of TANK 12"
   Circle "Circle_3" at 340,212 size 14x14
      Appearance <- "20_TANKS_IP_DATA_RIO_06_FIRST_TANK_BWT_LEVEL_HIHI"
   TextField "Text field_125" at 295,212 size 51x14; Text 'LS425-6P'
   Polyline "Polyline_1" at 261,205 size 123x240
      Visibility <- "504_Tank Grouping_DB2020_RUN TANK 12"
   TextField "Text field_64" at 288,273 size 74x20; Text 'Tank - 6P'
   Bar "Bar_2" at 394,206 size 122x241; MinimumValue 0; MaximumValue 100
      ProcessValue <- "20_TANKS_IP_DATA_RIO_05_FIRST_TANK_BWT_LEVEL"
   Button "Button_44" at 406,396 size 100x25; TextOff 'DISABLED'
      on Release: function_efd93a16("Tank 5P Status", 168, 315, -1, 2, 1)
      Visibility <- "504_Tank Grouping_DB2020_GROUP of TANK 10"
   Circle "Circle_4" at 472,212 size 14x14
      Appearance <- "20_TANKS_IP_DATA_RIO_05_FIRST_TANK_BWT_LEVEL_HIHI"
   TextField "Text field_124" at 427,212 size 51x14; Text 'LS425-5P'
   Polyline "Polyline_2" at 392,205 size 123x240
      Visibility <- "504_Tank Grouping_DB2020_RUN TANK 10"
   TextField "Text field_8" at 418,275 size 74x20; Text 'Tank - 5P'
   Bar "Bar_3" at 525,206 size 122x241; MinimumValue 0; MaximumValue 100
      ProcessValue <- "20_TANKS_IP_DATA_RIO_04_FIRST_TANK_BWT_LEVEL"
   Button "Button_40" at 537,395 size 100x25; TextOff 'DISABLED'
      on Release: function_efd93a16("Tank 4P Status", 168, 315, -1, 2, 1)
      Visibility <- "504_Tank Grouping_DB2020_GROUP of TANK 8"
   Circle "Circle_5" at 604,212 size 14x14
      Appearance <- "20_TANKS_IP_DATA_RIO_04_FIRST_TANK_BWT_LEVEL_HIHI"
   TextField "Text field_123" at 559,212 size 51x14; Text 'LS425-4P'
   Polyline "Polyline_3" at 525,205 size 123x240
      Visibility <- "504_Tank Grouping_DB2020_RUN TANK 8"
   TextField "Text field_9" at 553,275 size 74x20; Text 'Tank - 4P'
   Bar "Bar_4" at 657,206 size 122x241; MinimumValue 0; MaximumValue 100
      ProcessValue <- "20_TANKS_IP_DATA_RIO_03_FIRST_TANK_BWT_LEVEL"
   Button "Button_36" at 668,395 size 100x25; TextOff 'DISABLED'
      on Release: function_efd93a16("Tank 3P Status", 168, 315, -1, 0, 1)
      Visibility <- "504_Tank Grouping_DB2020_GROUP of TANK 6"
   Circle "Circle_7" at 736,212 size 14x14
      Appearance <- "20_TANKS_IP_DATA_RIO_03_FIRST_TANK_BWT_LEVEL_HIHI"
   TextField "Text field_122" at 691,212 size 51x14; Text 'LS425-3P'
   Polyline "Polyline_4" at 656,205 size 123x240
      Visibility <- "504_Tank Grouping_DB2020_RUN TANK 6"
   TextField "Text field_14" at 680,275 size 74x20; Text 'Tank - 3P'
   Bar "Bar_5" at 789,206 size 122x241; MinimumValue 0; MaximumValue 100
      ProcessValue <- "20_TANKS_IP_DATA_RIO_02_FIRST_TANK_BWT_LEVEL"
   Button "Button_32" at 802,396 size 100x25; TextOff 'DISABLED'
      on Release: function_efd93a16("Tank 2P Status", 168, 315, -1, 0, 1)
      Visibility <- "504_Tank Grouping_DB2020_GROUP of TANK 4"
   Circle "Circle_15" at 868,212 size 14x14
      Appearance <- "20_TANKS_IP_DATA_RIO_02_FIRST_TANK_BWT_LEVEL_HIHI"
   TextField "Text field_121" at 823,212 size 51x14; Text 'LS425-2P'
   Polyline "Polyline_5" at 789,205 size 123x240
      Visibility <- "504_Tank Grouping_DB2020_RUN TANK 4"
   TextField "Text field_15" at 816,275 size 74x20; Text 'Tank - 2P'
   Bar "Bar_6" at 922,205 size 122x241; MinimumValue 0; MaximumValue 100
      ProcessValue <- "20_TANKS_IP_DATA_RIO_01_SECOND_TANK_BWT_LEVEL"
   Button "Button_52" at 934,395 size 100x25; TextOff 'DISABLED'
      on Release: function_efd93a16("Tank 1P Status", 168, 315, -1, 0, 1)
      Visibility <- "504_Tank Grouping_DB2020_GROUP of TANK 2"
   Circle "Circle_16" at 999,211 size 14x14
      Appearance <- "20_TANKS_IP_DATA_RIO_01_SECOND_TANK_BWT_LEVEL_HIHI"
   TextField "Text field_120" at 955,211 size 51x14; Text 'LS425-1P'
   Polyline "Polyline_6" at 921,205 size 123x240
      Visibility <- "504_Tank Grouping_DB2020_RUN TANK 2"
   GraphicView "Graphic view_6" at 127,446 size 591x12; Picture "Graphic_151"
   TextField "Text field_16" at 947,275 size 74x20; Text 'Tank - 1P'
   Bar "Bar_7" at 1096,334 size 122x241; MinimumValue 0; MaximumValue 100
      ProcessValue <- "20_TANKS_IP_DATA_RIO_01_FIRST_TANK_BWT_LEVEL"
   Circle "Circle_24" at 1168,339 size 14x14
      Appearance <- "20_TANKS_IP_DATA_RIO_01_FIRST_TANK_BWT_LEVEL_HIHI"
   TextField "Text field_133" at 1139,339 size 35x14; Text 'LS425'
   Polyline "Polyline_14" at 1095,332 size 125x242
      Visibility <- "504_Tank Grouping_DB2020_RUN TANK 1"
   Button "Button_56" at 1110,524 size 100x25; TextOff 'DISABLED'
      on Release: function_efd93a16("Tank FP Status", 168, 315, -1, 0, 1)
      Visibility <- "504_Tank Grouping_DB2020_GROUP of TANK 1"
   TextField "Text field_17" at 1111,400 size 111x20; Text 'Fore PeakTank'
   Bar "Bar_8" at 922,458 size 122x258; MinimumValue 0; MaximumValue 100
      ProcessValue <- "20_TANKS_IP_DATA_RIO_01_THIRD_TANK_BWT_LEVEL"
   Button "Button_54" at 933,661 size 100x25; TextOff 'DISABLED'
      on Release: function_efd93a16("Tank 1S Status", 168, 315, -1, 0, 1)
      Visibility <- "504_Tank Grouping_DB2020_GROUP of TANK 3"
   Circle "Circle_23" at 1000,464 size 14x14
      Appearance <- "20_TANKS_IP_DATA_RIO_01_THIRD_TANK_BWT_LEVEL_HIHI"
   TextField "Text field_126" at 955,465 size 51x14; Text 'LS422-1S'
   Polyline "Polyline_7" at 921,458 size 123x259
      Visibility <- "504_Tank Grouping_DB2020_RUN TANK 3"
   TextField "Text field_10" at 950,618 size 74x20; Text 'Tank - 1S'
   Bar "Bar_9" at 790,459 size 122x258; MinimumValue 0; MaximumValue 100
      ProcessValue <- "20_TANKS_IP_DATA_RIO_02_SECOND_TANK_BWT_LEVEL"
   Button "Button_34" at 801,662 size 100x25; TextOff 'DISABLED'
      on Release: function_efd93a16("Tank 2S Status", 168, 315, -1, 0, 1)
      Visibility <- "504_Tank Grouping_DB2020_GROUP of TANK 5"
   Circle "Circle_22" at 868,465 size 14x14
      Appearance <- "20_TANKS_IP_DATA_RIO_02_SECOND_TANK_BWT_LEVEL_HIHI"
   TextField "Text field_127" at 823,466 size 51x14; Text 'LS422-2S'
   Polyline "Polyline_8" at 789,458 size 123x259
      Visibility <- "504_Tank Grouping_DB2020_RUN TANK 5"
   TextField "Text field_11" at 817,618 size 74x20; Text 'Tank - 2S'
   Bar "Bar_10" at 659,460 size 122x258; MinimumValue 0; MaximumValue 100
      ProcessValue <- "20_TANKS_IP_DATA_RIO_03_SECOND_TANK_BWT_LEVEL"
   Button "Button_38" at 669,663 size 100x25; TextOff 'DISABLED'
      on Release: function_efd93a16("Tank 3S Status", 168, 315, -1, 0, 1)
      Visibility <- "504_Tank Grouping_DB2020_GROUP of TANK 7"
   Circle "Circle_21" at 736,467 size 14x14
      Appearance <- "20_TANKS_IP_DATA_RIO_03_SECOND_TANK_BWT_LEVEL_HIHI"
   TextField "Text field_128" at 691,468 size 51x14; Text 'LS422-3S'
   Polyline "Polyline_9" at 658,458 size 123x259
      Visibility <- "504_Tank Grouping_DB2020_RUN TANK 7"
   TextField "Text field_12" at 690,618 size 74x20; Text 'Tank - 3S'
   Bar "Bar_11" at 526,459 size 122x258; MinimumValue 0; MaximumValue 100
      ProcessValue <- "20_TANKS_IP_DATA_RIO_04_SECOND_TANK_BWT_LEVEL"
   Button "Button_42" at 537,662 size 100x25; TextOff 'DISABLED'
      on Release: function_efd93a16("Tank 4S Status", 168, 315, -1, 2, 1)
      Visibility <- "504_Tank Grouping_DB2020_GROUP of TANK 9"
   Circle "Circle_19" at 604,466 size 14x14
      Appearance <- "20_TANKS_IP_DATA_RIO_04_SECOND_TANK_BWT_LEVEL_HIHI"
   TextField "Text field_129" at 559,467 size 51x14; Text 'LS422-4S'
   Polyline "Polyline_10" at 525,458 size 123x259
      Visibility <- "504_Tank Grouping_DB2020_RUN TANK 9"
   TextField "Text field_13" at 554,618 size 74x20; Text 'Tank - 4S'
   Bar "Bar_12" at 394,459 size 122x258; MinimumValue 0; MaximumValue 100
      ProcessValue <- "20_TANKS_IP_DATA_RIO_05_SECOND_TANK_BWT_LEVEL"
   Button "Button_46" at 405,662 size 100x25; TextOff 'DISABLED'
      on Release: function_efd93a16("Tank 5S Status", 168, 315, -1, 2, 1)
      Visibility <- "504_Tank Grouping_DB2020_GROUP of TANK 11"
   Circle "Circle_18" at 472,465 size 14x14
      Appearance <- "20_TANKS_IP_DATA_RIO_05_SECOND_TANK_BWT_LEVEL_HIHI"
   TextField "Text field_130" at 427,466 size 51x14; Text 'LS422-5S'
   Polyline "Polyline_11" at 393,458 size 123x259
      Visibility <- "504_Tank Grouping_DB2020_RUN TANK 11"
   TextField "Text field_18" at 424,618 size 74x20; Text 'Tank - 5S'
   Bar "Bar_13" at 262,460 size 122x258; MinimumValue 0; MaximumValue 100
      ProcessValue <- "20_TANKS_IP_DATA_RIO_06_SECOND_TANK_BWT_LEVEL"
   Button "Button_50" at 273,663 size 100x25; TextOff 'DISABLED'
      on Release: function_efd93a16("Tank 6S Status", 168, 315, -1, 2, 1)
      Visibility <- "504_Tank Grouping_DB2020_GROUP of TANK 13"
   Circle "Circle_17" at 340,467 size 14x14
      Appearance <- "20_TANKS_IP_DATA_RIO_06_SECOND_TANK_BWT_LEVEL_HIHI"
   TextField "Text field_131" at 295,468 size 51x14; Text 'LS422-6S'
   Polyline "Polyline_12" at 261,458 size 123x258
      Visibility <- "504_Tank Grouping_DB2020_RUN TANK 13"
   TextField "Text field_19" at 290,618 size 74x20; Text 'Tank - 6S'
   Bar "Bar_14" at 39,324 size 119x258; Unit %; MinimumValue 0; MaximumValue 100
      ProcessValue <- "20_TANKS_IP_DATA_RIO_07_FIRST_TANK_BWT_LEVEL"
   Circle "Circle_25" at 108,330 size 14x14
      Appearance <- "20_TANKS_IP_DATA_RIO_07_FIRST_TANK_BWT_LEVEL_HIHI"
   TextField "Text field_132" at 79,330 size 35x14; Text 'LS425'
   Polyline "Polyline_13" at 38,324 size 121x259
      Visibility <- "504_Tank Grouping_DB2020_RUN TANK 14"
   Button "Button_58" at 48,527 size 100x25; TextOff 'DISABLED'
      on Release: function_efd93a16("Tank AP Status", 168, 315, -1, 2, 1)
      Visibility <- "504_Tank Grouping_DB2020_GROUP of TANK 14"
   Button "HmiScreenItemData_6" at 1043,144 size 116x50; TextOn 'Back'; TextOff 'Tank Status'
      on Release: ActivateScreen("Balast Water Treatment Plant", 0)
   Button "Button_2" at 252,437 size 37x30; TextOff 'DB&B'
      on Release: function_efd93a16("Double Block & Bleed Valve Monitoring", 250, 250, -1, -1, 1)
      Appearance <- "10_DI_DATA_CV407_OPN"
   TextField "Text field_65" at 190,398 size 46x25; Text 'PGC'
   TextField "Text field_75" at 183,480 size 60x20; Text 'Disabled'
   TextField "Text field_76" at 183,480 size 60x20; Text 'Enabled'
      Visibility <- "10_DI_DATA_E_400_RUN"
   GraphicView "Graphic view_76" at 185,421 size 57x55; Picture "Graphic_251"
   Button "Button_6" at 179,402 size 70x105; TextOff 'Text'
      on Release: ActivateScreen("PGC System", 0)
   TextField "Text field_20" at 53,396 size 103x20; Text 'Aft PeakTank'
   GraphicView "Graphic view_108" at 4,683 size 96x48; Picture "Left Arow"
   Button "HmiScreenItemData_14" at 3,660 size 106x93; TextOn 'Back'; TextOff 'Text'
      on Press: ActivateScreen("Inert Gas Conditioning Plant", 0)
   IOField "I/O field_1" at 68,460 size 84x25; FormatPattern 99.99; Unit m
      ProcessValue <- "Data_From_WBT_Level_APT m"
   IOField "I/O field_2" at 285,331 size 84x25; FormatPattern 99.99; Unit m
      ProcessValue <- "Data_From_WBT_Level_WBT_6P m"
   IOField "I/O field_3" at 418,331 size 84x25; FormatPattern 99.99; Unit m
      ProcessValue <- "Data_From_WBT_Level_WBT_5P m"
   IOField "I/O field_4" at 550,331 size 84x25; FormatPattern 99.99; Unit m
      ProcessValue <- "Data_From_WBT_Level_WBT_4P m"
   IOField "I/O field_5" at 681,331 size 84x25; FormatPattern 99.99; Unit m
      ProcessValue <- "Data_From_WBT_Level_WBT_3P m"
   IOField "I/O field_6" at 815,331 size 84x25; FormatPattern 99.99; Unit m
      ProcessValue <- "Data_From_WBT_Level_WBT_2P m"
   IOField "I/O field_7" at 949,331 size 84x25; FormatPattern 99.99; Unit m
      ProcessValue <- "Data_From_WBT_Level_WBT_1P m"
   IOField "I/O field_8" at 1124,459 size 84x25; FormatPattern 99.99; Unit m
      ProcessValue <- "Data_From_WBT_Level_FPT m"
   IOField "I/O field_9" at 945,555 size 84x25; FormatPattern 99.99; Unit m
      ProcessValue <- "Data_From_WBT_Level_WBT_1S m"
   IOField "I/O field_10" at 816,556 size 84x25; FormatPattern 99.99; Unit m
      ProcessValue <- "Data_From_WBT_Level_WBT_2S m"
   IOField "I/O field_11" at 685,558 size 84x25; FormatPattern 99.99; Unit m
      ProcessValue <- "Data_From_WBT_Level_WBT_3S m"
   IOField "I/O field_12" at 553,557 size 84x25; FormatPattern 99.99; Unit m
      ProcessValue <- "Data_From_WBT_Level_WBT_4S m"
   IOField "I/O field_13" at 418,558 size 84x25; FormatPattern 99.99; Unit m
      ProcessValue <- "Data_From_WBT_Level_WBT_5S m"
   IOField "I/O field_14" at 287,559 size 84x25; FormatPattern 99.99; Unit m
      ProcessValue <- "Data_From_WBT_Level_WBT_6S m"
   Button "Button_88" at 34,324 size 127x264; TextOff 'Text'
      on Release: function_efd93a16("Tank AP Status", 168, 315, -1, 0, 1)
      Appearance <- "504_Tank Grouping_DB2020_RUN TANK 14"
   Button "Button_86" at 259,458 size 126x260; TextOff 'Text'
      on Release: function_efd93a16("Tank 6S Status", 168, 315, -1, 0, 1)
      Appearance <- "504_Tank Grouping_DB2020_RUN TANK 13"
   Button "Button_79" at 391,457 size 126x262; TextOff 'Text'
      on Release: function_efd93a16("Tank 5S Status", 168, 315, -1, 0, 1)
      Appearance <- "504_Tank Grouping_DB2020_RUN TANK 11"
   Button "Button_77" at 523,457 size 126x262; TextOff 'Text'
      on Release: function_efd93a16("Tank 4S Status", 168, 315, -1, 0, 1)
      Appearance <- "504_Tank Grouping_DB2020_RUN TANK 9"
   Button "Button_74" at 657,457 size 126x262; TextOff 'Text'
      on Release: function_efd93a16("Tank 3S Status", 168, 315, -1, 0, 1)
      Appearance <- "504_Tank Grouping_DB2020_RUN TANK 7"